   2132: 'Carrier 33 Drive: Error internal communications', class No Acknowledgement, trigger "DB302_HMI_Faults_Carrier33_Faults_1" bit 3
   2133: 'Carrier 33 Drive: Motor overtemperature', class No Acknowledgement, trigger "DB302_HMI_Faults_Carrier33_Faults_1" bit 4
   2134: 'Carrier 33 Drive: Motor overcurrent', class No Acknowledgement, trigger "DB302_HMI_Faults_Carrier33_Faults_1" bit 5
   2135: 'Carrier 33 Drive: Infeed or power unit not ready', class No Acknowledgement, trigger "DB302_HMI_Faults_Carrier33_Faults_1" bit 6
   2136: 'Carrier 33 Drive: Short-circuit/ground fault detected', class No Acknowledgement, trigger "DB302_HMI_Faults_Carrier33_Faults_1" bit 7
   2137: 'Carrier 33 Drive: PROFINET Setpoint timeout', class No Acknowledgement, trigger "DB302_HMI_Faults_Carrier33_Faults_1" bit 8
   2138: 'Carrier 33 Power unit: Overcurrent', class No Acknowledgement, trigger "DB302_HMI_Faults_Carrier33_Faults_1" bit 9
   2139: 'Carrier 33 Power unit: DC link voltage overvoltage', class No Acknowledgement, trigger "DB302_HMI_Faults_Carrier33_Faults_1" bit 10
   2140: 'Carrier 33 Power unit: DC link voltage undervoltage', class No Acknowledgement, trigger "DB302_HMI_Faults_Carrier33_Faults_1" bit 11
   2141: 'Carrier 33 Power unit: Line phase failure in main circuit', class No Acknowledgement, trigger "DB302_HMI_Faults_Carrier33_Faults_1" bit 12
   2142: 'Carrier 33 Power unit: Phase failure motor cable', class No Acknowledgement, trigger "DB302_HMI_Faults_Carrier33_Faults_1" bit 13
   2143: 'Carrier 33 Power unit: Ground fault', class No Acknowledgement, trigger "DB302_HMI_Faults_Carrier33_Faults_1" bit 14
   2144: 'Spare_Fault_2144', class No Acknowledgement, trigger "DB302_HMI_Faults_Carrier33_Faults_1" bit 15
   2145: 'Carrier 33 Motion Off Fault', class No Acknowledgement, trigger "DB302_HMI_Faults_Carrier33_Faults_2" bit 0
   2146: 'Carrier 33 Motion On Fault', class No Acknowledgement, trigger "DB302_HMI_Faults_Carrier33_Faults_2" bit 1
   2147: 'Carrier 33 Spacing Fault', class No Acknowledgement, trigger "DB302_HMI_Faults_Carrier33_Faults_2" bit 2
   2148: 'Carrier 33 Duplicate Carrier Number Fault', class No Acknowledgement, trigger "DB302_HMI_Faults_Carrier33_Faults_2" bit 3
   2149: 'Spare_Fault_2149', class No Acknowledgement, trigger "DB302_HMI_Faults_Carrier33_Faults_2" bit 4
   2150: 'Spare_Fault_2150', class No Acknowledgement, trigger "DB302_HMI_Faults_Carrier33_Faults_2" bit 5
   2151: 'Spare_Fault_2151', class No Acknowledgement, trigger "DB302_HMI_Faults_Carrier33_Faults_2" bit 6
   2152: 'Spare_Fault_2152', class No Acknowledgement, trigger "DB302_HMI_Faults_Carrier33_Faults_2" bit 7
   2153: 'Spare_Fault_2153', class No Acknowledgement, trigger "DB302_HMI_Faults_Carrier33_Faults_2" bit 8
   2154: 'Spare_Fault_2154', class No Acknowledgement, trigger "DB302_HMI_Faults_Carrier33_Faults_2" bit 9
   2155: 'Spare_Fault_2155', class No Acknowledgement, trigger "DB302_HMI_Faults_Carrier33_Faults_2" bit 10
   2156: 'Spare_Fault_2156', class No Acknowledgement, trigger "DB302_HMI_Faults_Carrier33_Faults_2" bit 11
   2157: 'Spare_Fault_2157', class No Acknowledgement, trigger "DB302_HMI_Faults_Carrier33_Faults_2" bit 12
   2158: 'Spare_Fault_2158', class No Acknowledgement, trigger "DB302_HMI_Faults_Carrier33_Faults_2" bit 13
   2159: 'Spare_Fault_2159', class No Acknowledgement, trigger "DB302_HMI_Faults_Carrier33_Faults_2" bit 14
   2160: 'Spare_Fault_2160', class No Acknowledgement, trigger "DB302_HMI_Faults_Carrier33_Faults_2" bit 15
   2161: 'Spare_Fault_2161', class No Acknowledgement, trigger "DB302_HMI_Faults_Carrier33_Faults_3" bit 0
   2162: 'Spare_Fault_2162', class No Acknowledgement, trigger "DB302_HMI_Faults_Carrier33_Faults_3" bit 1
   2163: 'Spare_Fault_2163', class No Acknowledgement, trigger "DB302_HMI_Faults_Carrier33_Faults_3" bit 2
   2164: 'Spare_Fault_2164', class No Acknowledgement, trigger "DB302_HMI_Faults_Carrier33_Faults_3" bit 3
   2165: 'Spare_Fault_2165', class No Acknowledgement, trigger "DB302_HMI_Faults_Carrier33_Faults_3" bit 4
   2166: 'Spare_Fault_2166', class No Acknowledgement, trigger "DB302_HMI_Faults_Carrier33_Faults_3" bit 5
   2167: 'Spare_Fault_2167', class No Acknowledgement, trigger "DB302_HMI_Faults_Carrier33_Faults_3" bit 6
   2168: 'Spare_Fault_2168', class No Acknowledgement, trigger "DB302_HMI_Faults_Carrier33_Faults_3" bit 7
   2169: 'Spare_Fault_2169', class No Acknowledgement, trigger "DB302_HMI_Faults_Carrier33_Faults_3" bit 8
   2170: 'Spare_Fault_2170', class No Acknowledgement, trigger "DB302_HMI_Faults_Carrier33_Faults_3" bit 9
   2171: 'Spare_Fault_2171', class No Acknowledgement, trigger "DB302_HMI_Faults_Carrier33_Faults_3" bit 10
   2172: 'Spare_Fault_2172', class No Acknowledgement, trigger "DB302_HMI_Faults_Carrier33_Faults_3" bit 11
   2173: 'Spare_Fault_2173', class No Acknowledgement, trigger "DB302_HMI_Faults_Carrier33_Faults_3" bit 12
   2174: 'Spare_Fault_2174', class No Acknowledgement, trigger "DB302_HMI_Faults_Carrier33_Faults_3" bit 13
   2175: 'Spare_Fault_2175', class No Acknowledgement, trigger "DB302_HMI_Faults_Carrier33_Faults_3" bit 14
   2176: 'Spare_Fault_2176', class No Acknowledgement, trigger "DB302_HMI_Faults_Carrier33_Faults_3" bit 15
   2177: 'Carrier 34 Disconnect Open Power Fault DI11.0', class No Acknowledgement, trigger "DB302_HMI_Faults_Carrier34_Faults_0" bit 0
   2178: 'Carrier 34 Drive Profinet Comm Fault', class No Acknowledgement, trigger "DB302_HMI_Faults_Carrier34_Faults_0" bit 1
   2179: 'Carrier 34 Production Stop Not Reset', class No Acknowledgement, trigger "DB302_HMI_Faults_Carrier34_Faults_0" bit 2
   2180: 'Carrier 34 CB02122 Tripped', class No Acknowledgement, trigger "DB302_HMI_Faults_Carrier34_Faults_0" bit 3
   2181: 'Carrier 34 CB02123 Tripped', class No Acknowledgement, trigger "DB302_HMI_Faults_Carrier34_Faults_0" bit 4
   2182: 'Carrier 34 AUX1 CB Tripped', class No Acknowledgement, trigger "DB302_HMI_Faults_Carrier34_Faults_0" bit 5
   2183: 'Carrier 34 AUX2 CB Tripped', class No Acknowledgement, trigger "DB302_HMI_Faults_Carrier34_Faults_0" bit 6
   2184: 'Carrier 34 PLC Not Communicating', class No Acknowledgement, trigger "DB302_HMI_Faults_Carrier34_Faults_0" bit 7
   2185: 'Carrier 34 Safe Input Card Fault', class No Acknowledgement, trigger "DB302_HMI_Faults_Carrier34_Faults_0" bit 8
   2186: 'Carrier 34 Safe Output Card Fault', class No Acknowledgement, trigger "DB302_HMI_Faults_Carrier34_Faults_0" bit 9
   2187: 'Carrier 34 Standard Input Card Fault', class No Acknowledgement, trigger "DB302_HMI_Faults_Carrier34_Faults_0" bit 10
   2188: 'Carrier 34 Standard Output Card Fault', class No Acknowledgement, trigger "DB302_HMI_Faults_Carrier34_Faults_0" bit 11
   2189: 'Carrier 34 Encoder Position Fault', class No Acknowledgement, trigger "DB302_HMI_Faults_Carrier34_Faults_0" bit 12
   2190: 'Carrier 34 Encoder Internal Error', class No Acknowledgement, trigger "DB302_HMI_Faults_Carrier34_Faults_0" bit 13
   2191: 'Carrier 34 Encoder Comm Fault', class No Acknowledgement, trigger "DB302_HMI_Faults_Carrier34_Faults_0" bit 14
   2192: 'Carrier 34 HMI Comm Fault', class No Acknowledgement, trigger "DB302_HMI_Faults_Carrier34_Faults_0" bit 15
   2193: 'Carrier 34 Crash Detection Fault', class No Acknowledgement, trigger "DB302_HMI_Faults_Carrier34_Faults_1" bit 0
   2194: 'Carrier 34 Carrier Number Invalid', class No Acknowledgement, trigger "DB302_HMI_Faults_Carrier34_Faults_1" bit 1
   2195: 'Carrier 34 Drive: PROFINET configuration error', class No Acknowledgement, trigger "DB302_HMI_Faults_Carrier34_Faults_1" bit 2
   2196: 'Carrier 34 Drive: Error internal communications', class No Acknowledgement, trigger "DB302_HMI_Faults_Carrier34_Faults_1" bit 3
   2197: 'Carrier 34 Drive: Motor overtemperature', class No Acknowledgement, trigger "DB302_HMI_Faults_Carrier34_Faults_1" bit 4
   2198: 'Carrier 34 Drive: Motor overcurrent', class No Acknowledgement, trigger "DB302_HMI_Faults_Carrier34_Faults_1" bit 5
   2199: 'Carrier 34 Drive: Infeed or power unit not ready', class No Acknowledgement, trigger "DB302_HMI_Faults_Carrier34_Faults_1" bit 6
   2200: 'Carrier 34 Drive: Short-circuit/ground fault detected', class No Acknowledgement, trigger "DB302_HMI_Faults_Carrier34_Faults_1" bit 7
   2201: 'Carrier 34 Drive: PROFINET Setpoint timeout', class No Acknowledgement, trigger "DB302_HMI_Faults_Carrier34_Faults_1" bit 8
   2202: 'Carrier 34 Power unit: Overcurrent', class No Acknowledgement, trigger "DB302_HMI_Faults_Carrier34_Faults_1" bit 9
   2203: 'Carrier 34 Power unit: DC link voltage overvoltage', class No Acknowledgement, trigger "DB302_HMI_Faults_Carrier34_Faults_1" bit 10
   2204: 'Carrier 34 Power unit: DC link voltage undervoltage', class No Acknowledgement, trigger "DB302_HMI_Faults_Carrier34_Faults_1" bit 11
   2205: 'Carrier 34 Power unit: Line phase failure in main circuit', class No Acknowledgement, trigger "DB302_HMI_Faults_Carrier34_Faults_1" bit 12
   2206: 'Carrier 34 Power unit: Phase failure motor cable', class No Acknowledgement, trigger "DB302_HMI_Faults_Carrier34_Faults_1" bit 13
   2207: 'Carrier 34 Power unit: Ground fault', class No Acknowledgement, trigger "DB302_HMI_Faults_Carrier34_Faults_1" bit 14
   2208: 'Spare_Fault_2208', class No Acknowledgement, trigger "DB302_HMI_Faults_Carrier34_Faults_1" bit 15
   2209: 'Carrier 34 Motion Off Fault', class No Acknowledgement, trigger "DB302_HMI_Faults_Carrier34_Faults_2" bit 0
   2210: 'Carrier 34 Motion On Fault', class No Acknowledgement, trigger "DB302_HMI_Faults_Carrier34_Faults_2" bit 1
   2211: 'Carrier 34 Spacing Fault', class No Acknowledgement, trigger "DB302_HMI_Faults_Carrier34_Faults_2" bit 2
   2212: 'Carrier 34 Duplicate Carrier Number Fault', class No Acknowledgement, trigger "DB302_HMI_Faults_Carrier34_Faults_2" bit 3
   2213: 'Spare_Fault_2213', class No Acknowledgement, trigger "DB302_HMI_Faults_Carrier34_Faults_2" bit 4
   2214: 'Spare_Fault_2214', class No Acknowledgement, trigger "DB302_HMI_Faults_Carrier34_Faults_2" bit 5
   2215: 'Spare_Fault_2215', class No Acknowledgement, trigger "DB302_HMI_Faults_Carrier34_Faults_2" bit 6
   2216: 'Spare_Fault_2216', class No Acknowledgement, trigger "DB302_HMI_Faults_Carrier34_Faults_2" bit 7
   2217: 'Spare_Fault_2217', class No Acknowledgement, trigger "DB302_HMI_Faults_Carrier34_Faults_2" bit 8
   2218: 'Spare_Fault_2218', class No Acknowledgement, trigger "DB302_HMI_Faults_Carrier34_Faults_2" bit 9
   2219: 'Spare_Fault_2219', class No Acknowledgement, trigger "DB302_HMI_Faults_Carrier34_Faults_2" bit 10
   2220: 'Spare_Fault_2220', class No Acknowledgement, trigger "DB302_HMI_Faults_Carrier34_Faults_2" bit 11
   2221: 'Spare_Fault_2221', class No Acknowledgement, trigger "DB302_HMI_Faults_Carrier34_Faults_2" bit 12
   2222: 'Spare_Fault_2222', class No Acknowledgement, trigger "DB302_HMI_Faults_Carrier34_Faults_2" bit 13
   2223: 'Spare_Fault_2223', class No Acknowledgement, trigger "DB302_HMI_Faults_Carrier34_Faults_2" bit 14
   2224: 'Spare_Fault_2224', class No Acknowledgement, trigger "DB302_HMI_Faults_Carrier34_Faults_2" bit 15
   2225: 'Spare_Fault_2225', class No Acknowledgement, trigger "DB302_HMI_Faults_Carrier34_Faults_3" bit 0
   2226: 'Spare_Fault_2226', class No Acknowledgement, trigger "DB302_HMI_Faults_Carrier34_Faults_3" bit 1
   2227: 'Spare_Fault_2227', class No Acknowledgement, trigger "DB302_HMI_Faults_Carrier34_Faults_3" bit 2
   2228: 'Spare_Fault_2228', class No Acknowledgement, trigger "DB302_HMI_Faults_Carrier34_Faults_3" bit 3
   2229: 'Spare_Fault_2229', class No Acknowledgement, trigger "DB302_HMI_Faults_Carrier34_Faults_3" bit 4
   2230: 'Spare_Fault_2230', class No Acknowledgement, trigger "DB302_HMI_Faults_Carrier34_Faults_3" bit 5
   2231: 'Spare_Fault_2231', class No Acknowledgement, trigger "DB302_HMI_Faults_Carrier34_Faults_3" bit 6
   2232: 'Spare_Fault_2232', class No Acknowledgement, trigger "DB302_HMI_Faults_Carrier34_Faults_3" bit 7
   2233: 'Spare_Fault_2233', class No Acknowledgement, trigger "DB302_HMI_Faults_Carrier34_Faults_3" bit 8
   2234: 'Spare_Fault_2234', class No Acknowledgement, trigger "DB302_HMI_Faults_Carrier34_Faults_3" bit 9
   2235: 'Spare_Fault_2235', class No Acknowledgement, trigger "DB302_HMI_Faults_Carrier34_Faults_3" bit 10
   2236: 'Spare_Fault_2236', class No Acknowledgement, trigger "DB302_HMI_Faults_Carrier34_Faults_3" bit 11
   2237: 'Spare_Fault_2237', class No Acknowledgement, trigger "DB302_HMI_Faults_Carrier34_Faults_3" bit 12
   2238: 'Spare_Fault_2238', class No Acknowledgement, trigger "DB302_HMI_Faults_Carrier34_Faults_3" bit 13
   2239: 'Spare_Fault_2239', class No Acknowledgement, trigger "DB302_HMI_Faults_Carrier34_Faults_3" bit 14
   2240: 'Spare_Fault_2240', class No Acknowledgement, trigger "DB302_HMI_Faults_Carrier34_Faults_3" bit 15
   2241: 'Carrier 35 Disconnect Open Power Fault DI11.0', class No Acknowledgement, trigger "DB302_HMI_Faults_Carrier35_Faults_0" bit 0
   2242: 'Carrier 35 Drive Profinet Comm Fault', class No Acknowledgement, trigger "DB302_HMI_Faults_Carrier35_Faults_0" bit 1
   2243: 'Carrier 35 Production Stop Not Reset', class No Acknowledgement, trigger "DB302_HMI_Faults_Carrier35_Faults_0" bit 2
   2244: 'Carrier 35 CB02122 Tripped', class No Acknowledgement, trigger "DB302_HMI_Faults_Carrier35_Faults_0" bit 3
   2245: 'Carrier 35 CB02123 Tripped', class No Acknowledgement, trigger "DB302_HMI_Faults_Carrier35_Faults_0" bit 4
   2246: 'Carrier 35 AUX1 CB Tripped', class No Acknowledgement, trigger "DB302_HMI_Faults_Carrier35_Faults_0" bit 5
   2247: 'Carrier 35 AUX2 CB Tripped', class No Acknowledgement, trigger "DB302_HMI_Faults_Carrier35_Faults_0" bit 6
   2248: 'Carrier 35 PLC Not Communicating', class No Acknowledgement, trigger "DB302_HMI_Faults_Carrier35_Faults_0" bit 7
   2249: 'Carrier 35 Safe Input Card Fault', class No Acknowledgement, trigger "DB302_HMI_Faults_Carrier35_Faults_0" bit 8
   2250: 'Carrier 35 Safe Output Card Fault', class No Acknowledgement, trigger "DB302_HMI_Faults_Carrier35_Faults_0" bit 9
   2251: 'Carrier 35 Standard Input Card Fault', class No Acknowledgement, trigger "DB302_HMI_Faults_Carrier35_Faults_0" bit 10
   2252: 'Carrier 35 Standard Output Card Fault', class No Acknowledgement, trigger "DB302_HMI_Faults_Carrier35_Faults_0" bit 11
   2253: 'Carrier 35 Encoder Position Fault', class No Acknowledgement, trigger "DB302_HMI_Faults_Carrier35_Faults_0" bit 12
   2254: 'Carrier 35 Encoder Internal Error', class No Acknowledgement, trigger "DB302_HMI_Faults_Carrier35_Faults_0" bit 13
   2255: 'Carrier 35 Encoder Comm Fault', class No Acknowledgement, trigger "DB302_HMI_Faults_Carrier35_Faults_0" bit 14
   2256: 'Carrier 35 HMI Comm Fault', class No Acknowledgement, trigger "DB302_HMI_Faults_Carrier35_Faults_0" bit 15
   2257: 'Carrier 35 Crash Detection Fault', class No Acknowledgement, trigger "DB302_HMI_Faults_Carrier35_Faults_1" bit 0
   2258: 'Carrier 35 Carrier Number Invalid', class No Acknowledgement, trigger "DB302_HMI_Faults_Carrier35_Faults_1" bit 1
   2259: 'Carrier 35 Drive: PROFINET configuration error', class No Acknowledgement, trigger "DB302_HMI_Faults_Carrier35_Faults_1" bit 2
   2260: 'Carrier 35 Drive: Error internal communications', class No Acknowledgement, trigger "DB302_HMI_Faults_Carrier35_Faults_1" bit 3
   2261: 'Carrier 35 Drive: Motor overtemperature', class No Acknowledgement, trigger "DB302_HMI_Faults_Carrier35_Faults_1" bit 4
   2262: 'Carrier 35 Drive: Motor overcurrent', class No Acknowledgement, trigger "DB302_HMI_Faults_Carrier35_Faults_1" bit 5
   2263: 'Carrier 35 Drive: Infeed or power unit not ready', class No Acknowledgement, trigger "DB302_HMI_Faults_Carrier35_Faults_1" bit 6
   2264: 'Carrier 35 Drive: Short-circuit/ground fault detected', class No Acknowledgement, trigger "DB302_HMI_Faults_Carrier35_Faults_1" bit 7
   2265: 'Carrier 35 Drive: PROFINET Setpoint timeout', class No Acknowledgement, trigger "DB302_HMI_Faults_Carrier35_Faults_1" bit 8
   2266: 'Carrier 35 Power unit: Overcurrent', class No Acknowledgement, trigger "DB302_HMI_Faults_Carrier35_Faults_1" bit 9
   2267: 'Carrier 35 Power unit: DC link voltage overvoltage', class No Acknowledgement, trigger "DB302_HMI_Faults_Carrier35_Faults_1" bit 10
   2268: 'Carrier 35 Power unit: DC link voltage undervoltage', class No Acknowledgement, trigger "DB302_HMI_Faults_Carrier35_Faults_1" bit 11
   2269: 'Carrier 35 Power unit: Line phase failure in main circuit', class No Acknowledgement, trigger "DB302_HMI_Faults_Carrier35_Faults_1" bit 12
   2270: 'Carrier 35 Power unit: Phase failure motor cable', class No Acknowledgement, trigger "DB302_HMI_Faults_Carrier35_Faults_1" bit 13
   2271: 'Carrier 35 Power unit: Ground fault', class No Acknowledgement, trigger "DB302_HMI_Faults_Carrier35_Faults_1" bit 14
   2272: 'Spare_Fault_2272', class No Acknowledgement, trigger "DB302_HMI_Faults_Carrier35_Faults_1" bit 15
   2273: 'Carrier 35 Motion Off Fault', class No Acknowledgement, trigger "DB302_HMI_Faults_Carrier35_Faults_2" bit 0
   2274: 'Carrier 35 Motion On Fault', class No Acknowledgement, trigger "DB302_HMI_Faults_Carrier35_Faults_2" bit 1
   2275: 'Carrier 35 Spacing Fault', class No Acknowledgement, trigger "DB302_HMI_Faults_Carrier35_Faults_2" bit 2
   2276: 'Carrier 35 Duplicate Carrier Number Fault', class No Acknowledgement, trigger "DB302_HMI_Faults_Carrier35_Faults_2" bit 3
   2277: 'Spare_Fault_2277', class No Acknowledgement, trigger "DB302_HMI_Faults_Carrier35_Faults_2" bit 4
   2278: 'Spare_Fault_2278', class No Acknowledgement, trigger "DB302_HMI_Faults_Carrier35_Faults_2" bit 5
   2279: 'Spare_Fault_2279', class No Acknowledgement, trigger "DB302_HMI_Faults_Carrier35_Faults_2" bit 6
   2280: 'Spare_Fault_2280', class No Acknowledgement, trigger "DB302_HMI_Faults_Carrier35_Faults_2" bit 7
   2281: 'Spare_Fault_2281', class No Acknowledgement, trigger "DB302_HMI_Faults_Carrier35_Faults_2" bit 8
   2282: 'Spare_Fault_2282', class No Acknowledgement, trigger "DB302_HMI_Faults_Carrier35_Faults_2" bit 9
   2283: 'Spare_Fault_2283', class No Acknowledgement, trigger "DB302_HMI_Faults_Carrier35_Faults_2" bit 10
   2284: 'Spare_Fault_2284', class No Acknowledgement, trigger "DB302_HMI_Faults_Carrier35_Faults_2" bit 11
   2285: 'Spare_Fault_2285', class No Acknowledgement, trigger "DB302_HMI_Faults_Carrier35_Faults_2" bit 12
   2286: 'Spare_Fault_2286', class No Acknowledgement, trigger "DB302_HMI_Faults_Carrier35_Faults_2" bit 13
   2287: 'Spare_Fault_2287', class No Acknowledgement, trigger "DB302_HMI_Faults_Carrier35_Faults_2" bit 14
   2288: 'Spare_Fault_2288', class No Acknowledgement, trigger "DB302_HMI_Faults_Carrier35_Faults_2" bit 15
   2289: 'Spare_Fault_2289', class No Acknowledgement, trigger "DB302_HMI_Faults_Carrier35_Faults_3" bit 0
   2290: 'Spare_Fault_2290', class No Acknowledgement, trigger "DB302_HMI_Faults_Carrier35_Faults_3" bit 1
   2291: 'Spare_Fault_2291', class No Acknowledgement, trigger "DB302_HMI_Faults_Carrier35_Faults_3" bit 2
   2292: 'Spare_Fault_2292', class No Acknowledgement, trigger "DB302_HMI_Faults_Carrier35_Faults_3" bit 3
   2293: 'Spare_Fault_2293', class No Acknowledgement, trigger "DB302_HMI_Faults_Carrier35_Faults_3" bit 4
   2294: 'Spare_Fault_2294', class No Acknowledgement, trigger "DB302_HMI_Faults_Carrier35_Faults_3" bit 5
   2295: 'Spare_Fault_2295', class No Acknowledgement, trigger "DB302_HMI_Faults_Carrier35_Faults_3" bit 6
   2296: 'Spare_Fault_2296', class No Acknowledgement, trigger "DB302_HMI_Faults_Carrier35_Faults_3" bit 7
   2297: 'Spare_Fault_2297', class No Acknowledgement, trigger "DB302_HMI_Faults_Carrier35_Faults_3" bit 8
   2298: 'Spare_Fault_2298', class No Acknowledgement, trigger "DB302_HMI_Faults_Carrier35_Faults_3" bit 9
   2299: 'Spare_Fault_2299', class No Acknowledgement, trigger "DB302_HMI_Faults_Carrier35_Faults_3" bit 10
   2300: 'Spare_Fault_2300', class No Acknowledgement, trigger "DB302_HMI_Faults_Carrier35_Faults_3" bit 11
   2301: 'Spare_Fault_2301', class No Acknowledgement, trigger "DB302_HMI_Faults_Carrier35_Faults_3" bit 12
   2302: 'Spare_Fault_2302', class No Acknowledgement, trigger "DB302_HMI_Faults_Carrier35_Faults_3" bit 13
   2303: 'Spare_Fault_2303', class No Acknowledgement, trigger "DB302_HMI_Faults_Carrier35_Faults_3" bit 14
   2304: 'Spare_Fault_2304', class No Acknowledgement, trigger "DB302_HMI_Faults_Carrier35_Faults_3" bit 15
   2305: 'Carrier36 Disconnect Open Power Fault DI11.0', class No Acknowledgement, trigger "DB302_HMI_Faults_Carrier36_Faults_0" bit 0
   2306: 'Carrier36 Drive Profinet Comm Fault', class No Acknowledgement, trigger "DB302_HMI_Faults_Carrier36_Faults_0" bit 1
   2307: 'Carrier36 Production Stop Not Reset', class No Acknowledgement, trigger "DB302_HMI_Faults_Carrier36_Faults_0" bit 2
   2308: 'Carrier36 CB02122 Tripped', class No Acknowledgement, trigger "DB302_HMI_Faults_Carrier36_Faults_0" bit 3
   2309: 'Carrier36 CB02123 Tripped', class No Acknowledgement, trigger "DB302_HMI_Faults_Carrier36_Faults_0" bit 4
   2310: 'Carrier36 AUX1 CB Tripped', class No Acknowledgement, trigger "DB302_HMI_Faults_Carrier36_Faults_0" bit 5
   2311: 'Carrier36 AUX2 CB Tripped', class No Acknowledgement, trigger "DB302_HMI_Faults_Carrier36_Faults_0" bit 6
   2312: 'Carrier36 PLC Not Communicating', class No Acknowledgement, trigger "DB302_HMI_Faults_Carrier36_Faults_0" bit 7
   2313: 'Carrier36 Safe Input Card Fault', class No Acknowledgement, trigger "DB302_HMI_Faults_Carrier36_Faults_0" bit 8
   2314: 'Carrier36 Safe Output Card Fault', class No Acknowledgement, trigger "DB302_HMI_Faults_Carrier36_Faults_0" bit 9
   2315: 'Carrier36 Standard Input Card Fault', class No Acknowledgement, trigger "DB302_HMI_Faults_Carrier36_Faults_0" bit 10
   2316: 'Carrier36 Standard Output Card Fault', class No Acknowledgement, trigger "DB302_HMI_Faults_Carrier36_Faults_0" bit 11
   2317: 'Carrier36 Encoder Position Fault', class No Acknowledgement, trigger "DB302_HMI_Faults_Carrier36_Faults_0" bit 12
   2318: 'Carrier36 Encoder Internal Error', class No Acknowledgement, trigger "DB302_HMI_Faults_Carrier36_Faults_0" bit 13
   2319: 'Carrier36 Encoder Comm Fault', class No Acknowledgement, trigger "DB302_HMI_Faults_Carrier36_Faults_0" bit 14
   2320: 'Carrier36 HMI Comm Fault', class No Acknowledgement, trigger "DB302_HMI_Faults_Carrier36_Faults_0" bit 15
   2321: 'Carrier36 Crash Detection Fault', class No Acknowledgement, trigger "DB302_HMI_Faults_Carrier36_Faults_1" bit 0
   2322: 'Carrier36 Carrier Number Invalid', class No Acknowledgement, trigger "DB302_HMI_Faults_Carrier36_Faults_1" bit 1
   2323: 'Carrier36 Drive: PROFINET configuration error', class No Acknowledgement, trigger "DB302_HMI_Faults_Carrier36_Faults_1" bit 2
   2324: 'Carrier36 Drive: Error internal communications', class No Acknowledgement, trigger "DB302_HMI_Faults_Carrier36_Faults_1" bit 3
   2325: 'Carrier36 Drive: Motor overtemperature', class No Acknowledgement, trigger "DB302_HMI_Faults_Carrier36_Faults_1" bit 4
   2326: 'Carrier36 Drive: Motor overcurrent', class No Acknowledgement, trigger "DB302_HMI_Faults_Carrier36_Faults_1" bit 5
   2327: 'Carrier36 Drive: Infeed or power unit not ready', class No Acknowledgement, trigger "DB302_HMI_Faults_Carrier36_Faults_1" bit 6
   2328: 'Carrier36 Drive: Short-circuit/ground fault detected', class No Acknowledgement, trigger "DB302_HMI_Faults_Carrier36_Faults_1" bit 7
   2329: 'Carrier36 Drive: PROFINET Setpoint timeout', class No Acknowledgement, trigger "DB302_HMI_Faults_Carrier36_Faults_1" bit 8
   2330: 'Carrier36 Power unit: Overcurrent', class No Acknowledgement, trigger "DB302_HMI_Faults_Carrier36_Faults_1" bit 9
   2331: 'Carrier36 Power unit: DC link voltage overvoltage', class No Acknowledgement, trigger "DB302_HMI_Faults_Carrier36_Faults_1" bit 10
   2332: 'Carrier36 Power unit: DC link voltage undervoltage', class No Acknowledgement, trigger "DB302_HMI_Faults_Carrier36_Faults_1" bit 11
   2333: 'Carrier36 Power unit: Line phase failure in main circuit', class No Acknowledgement, trigger "DB302_HMI_Faults_Carrier36_Faults_1" bit 12
   2334: 'Carrier36 Power unit: Phase failure motor cable', class No Acknowledgement, trigger "DB302_HMI_Faults_Carrier36_Faults_1" bit 13
   2335: 'Carrier36 Power unit: Ground fault', class No Acknowledgement, trigger "DB302_HMI_Faults_Carrier36_Faults_1" bit 14
   2336: 'Spare_Fault_2336', class No Acknowledgement, trigger "DB302_HMI_Faults_Carrier36_Faults_1" bit 15
   2337: 'Carrier36 Motion Off Fault', class No Acknowledgement, trigger "DB302_HMI_Faults_Carrier36_Faults_2" bit 0
   2338: 'Carrier36 Motion On Fault', class No Acknowledgement, trigger "DB302_HMI_Faults_Carrier36_Faults_2" bit 1
   2339: 'Carrier36 Spacing Fault', class No Acknowledgement, trigger "DB302_HMI_Faults_Carrier36_Faults_2" bit 2
   2340: 'Carrier36 Duplicate Carrier Number Fault', class No Acknowledgement, trigger "DB302_HMI_Faults_Carrier36_Faults_2" bit 3
   2341: 'Spare_Fault_2341', class No Acknowledgement, trigger "DB302_HMI_Faults_Carrier36_Faults_2" bit 4
   2342: 'Spare_Fault_2342', class No Acknowledgement, trigger "DB302_HMI_Faults_Carrier36_Faults_2" bit 5
   2343: 'Spare_Fault_2343', class No Acknowledgement, trigger "DB302_HMI_Faults_Carrier36_Faults_2" bit 6
   2344: 'Spare_Fault_2344', class No Acknowledgement, trigger "DB302_HMI_Faults_Carrier36_Faults_2" bit 7
   2345: 'Spare_Fault_2345', class No Acknowledgement, trigger "DB302_HMI_Faults_Carrier36_Faults_2" bit 8
   2346: 'Spare_Fault_2346', class No Acknowledgement, trigger "DB302_HMI_Faults_Carrier36_Faults_2" bit 9
   2347: 'Spare_Fault_2347', class No Acknowledgement, trigger "DB302_HMI_Faults_Carrier36_Faults_2" bit 10
   2348: 'Spare_Fault_2348', class No Acknowledgement, trigger "DB302_HMI_Faults_Carrier36_Faults_2" bit 11
   2349: 'Spare_Fault_2349', class No Acknowledgement, trigger "DB302_HMI_Faults_Carrier36_Faults_2" bit 12
   2350: 'Spare_Fault_2350', class No Acknowledgement, trigger "DB302_HMI_Faults_Carrier36_Faults_2" bit 13
   2351: 'Spare_Fault_2351', class No Acknowledgement, trigger "DB302_HMI_Faults_Carrier36_Faults_2" bit 14
   2352: 'Spare_Fault_2352', class No Acknowledgement, trigger "DB302_HMI_Faults_Carrier36_Faults_2" bit 15
   2353: 'Spare_Fault_2353', class No Acknowledgement, trigger "DB302_HMI_Faults_Carrier36_Faults_3" bit 0
   2354: 'Spare_Fault_2354', class No Acknowledgement, trigger "DB302_HMI_Faults_Carrier36_Faults_3" bit 1
   2355: 'Spare_Fault_2355', class No Acknowledgement, trigger "DB302_HMI_Faults_Carrier36_Faults_3" bit 2
   2356: 'Spare_Fault_2356', class No Acknowledgement, trigger "DB302_HMI_Faults_Carrier36_Faults_3" bit 3
   2357: 'Spare_Fault_2357', class No Acknowledgement, trigger "DB302_HMI_Faults_Carrier36_Faults_3" bit 4
   2358: 'Spare_Fault_2358', class No Acknowledgement, trigger "DB302_HMI_Faults_Carrier36_Faults_3" bit 5
   2359: 'Spare_Fault_2359', class No Acknowledgement, trigger "DB302_HMI_Faults_Carrier36_Faults_3" bit 6
   2360: 'Spare_Fault_2360', class No Acknowledgement, trigger "DB302_HMI_Faults_Carrier36_Faults_3" bit 7
   2361: 'Spare_Fault_2361', class No Acknowledgement, trigger "DB302_HMI_Faults_Carrier36_Faults_3" bit 8
   2362: 'Spare_Fault_2362', class No Acknowledgement, trigger "DB302_HMI_Faults_Carrier36_Faults_3" bit 9
   2363: 'Spare_Fault_2363', class No Acknowledgement, trigger "DB302_HMI_Faults_Carrier36_Faults_3" bit 10
   2364: 'Spare_Fault_2364', class No Acknowledgement, trigger "DB302_HMI_Faults_Carrier36_Faults_3" bit 11
   2365: 'Spare_Fault_2365', class No Acknowledgement, trigger "DB302_HMI_Faults_Carrier36_Faults_3" bit 12
   2366: 'Spare_Fault_2366', class No Acknowledgement, trigger "DB302_HMI_Faults_Carrier36_Faults_3" bit 13
   2367: 'Spare_Fault_2367', class No Acknowledgement, trigger "DB302_HMI_Faults_Carrier36_Faults_3" bit 14
   2368: 'Spare_Fault_2368', class No Acknowledgement, trigger "DB302_HMI_Faults_Carrier36_Faults_3" bit 15
   2369: 'Carrier 37 Disconnect Open Power Fault DI11.0', class No Acknowledgement, trigger "DB302_HMI_Faults_Carrier37_Faults_0" bit 0
   2370: 'Carrier 37 Drive Profinet Comm Fault', class No Acknowledgement, trigger "DB302_HMI_Faults_Carrier37_Faults_0" bit 1
   2371: 'Carrier 37 Production Stop Not Reset', class No Acknowledgement, trigger "DB302_HMI_Faults_Carrier37_Faults_0" bit 2
   2372: 'Carrier 37 CB02122 Tripped', class No Acknowledgement, trigger "DB302_HMI_Faults_Carrier37_Faults_0" bit 3
   2373: 'Carrier 37 CB02123 Tripped', class No Acknowledgement, trigger "DB302_HMI_Faults_Carrier37_Faults_0" bit 4
   2374: 'Carrier 37 AUX1 CB Tripped', class No Acknowledgement, trigger "DB302_HMI_Faults_Carrier37_Faults_0" bit 5
   2375: 'Carrier 37 AUX2 CB Tripped', class No Acknowledgement, trigger "DB302_HMI_Faults_Carrier37_Faults_0" bit 6
   2376: 'Carrier 37 PLC Not Communicating', class No Acknowledgement, trigger "DB302_HMI_Faults_Carrier37_Faults_0" bit 7
   2377: 'Carrier 37 Safe Input Card Fault', class No Acknowledgement, trigger "DB302_HMI_Faults_Carrier37_Faults_0" bit 8
   2378: 'Carrier 37 Safe Output Card Fault', class No Acknowledgement, trigger "DB302_HMI_Faults_Carrier37_Faults_0" bit 9
   2379: 'Carrier 37 Standard Input Card Fault', class No Acknowledgement, trigger "DB302_HMI_Faults_Carrier37_Faults_0" bit 10
   2380: 'Carrier 37 Standard Output Card Fault', class No Acknowledgement, trigger "DB302_HMI_Faults_Carrier37_Faults_0" bit 11
   2381: 'Carrier 37 Encoder Position Fault', class No Acknowledgement, trigger "DB302_HMI_Faults_Carrier37_Faults_0" bit 12
   2382: 'Carrier 37 Encoder Internal Error', class No Acknowledgement, trigger "DB302_HMI_Faults_Carrier37_Faults_0" bit 13
   2383: 'Carrier 37 Encoder Comm Fault', class No Acknowledgement, trigger "DB302_HMI_Faults_Carrier37_Faults_0" bit 14
   2384: 'Carrier 37 HMI Comm Fault', class No Acknowledgement, trigger "DB302_HMI_Faults_Carrier37_Faults_0" bit 15
   2385: 'Carrier 37 Crash Detection Fault', class No Acknowledgement, trigger "DB302_HMI_Faults_Carrier37_Faults_1" bit 0
   2386: 'Carrier 37 Carrier Number Invalid', class No Acknowledgement, trigger "DB302_HMI_Faults_Carrier37_Faults_1" bit 1
   2387: 'Carrier 37 Drive: PROFINET configuration error', class No Acknowledgement, trigger "DB302_HMI_Faults_Carrier37_Faults_1" bit 2
   2388: 'Carrier 37 Drive: Error internal communications', class No Acknowledgement, trigger "DB302_HMI_Faults_Carrier37_Faults_1" bit 3
   2389: 'Carrier 37 Drive: Motor overtemperature', class No Acknowledgement, trigger "DB302_HMI_Faults_Carrier37_Faults_1" bit 4
   2390: 'Carrier 37 Drive: Motor overcurrent', class No Acknowledgement, trigger "DB302_HMI_Faults_Carrier37_Faults_1" bit 5
   2391: 'Carrier 37 Drive: Infeed or power unit not ready', class No Acknowledgement, trigger "DB302_HMI_Faults_Carrier37_Faults_1" bit 6
   2392: 'Carrier 37 Drive: Short-circuit/ground fault detected', class No Acknowledgement, trigger "DB302_HMI_Faults_Carrier37_Faults_1" bit 7
   2393: 'Carrier 37 Drive: PROFINET Setpoint timeout', class No Acknowledgement, trigger "DB302_HMI_Faults_Carrier37_Faults_1" bit 8
   2394: 'Carrier 37 Power unit: Overcurrent', class No Acknowledgement, trigger "DB302_HMI_Faults_Carrier37_Faults_1" bit 9
   2395: 'Carrier 37 Power unit: DC link voltage overvoltage', class No Acknowledgement, trigger "DB302_HMI_Faults_Carrier37_Faults_1" bit 10
   2396: 'Carrier 37 Power unit: DC link voltage undervoltage', class No Acknowledgement, trigger "DB302_HMI_Faults_Carrier37_Faults_1" bit 11
   2397: 'Carrier 37 Power unit: Line phase failure in main circuit', class No Acknowledgement, trigger "DB302_HMI_Faults_Carrier37_Faults_1" bit 12
   2398: 'Carrier 37 Power unit: Phase failure motor cable', class No Acknowledgement, trigger "DB302_HMI_Faults_Carrier37_Faults_1" bit 13
   2399: 'Carrier 37 Power unit: Ground fault', class No Acknowledgement, trigger "DB302_HMI_Faults_Carrier37_Faults_1" bit 14
   2400: 'Spare_Fault_2400', class No Acknowledgement, trigger "DB302_HMI_Faults_Carrier37_Faults_1" bit 15
   2401: 'Carrier 37 Motion Off Fault', class No Acknowledgement, trigger "DB302_HMI_Faults_Carrier37_Faults_2" bit 0
   2402: 'Carrier 37 Motion On Fault', class No Acknowledgement, trigger "DB302_HMI_Faults_Carrier37_Faults_2" bit 1
   2403: 'Carrier 37 Spacing Fault', class No Acknowledgement, trigger "DB302_HMI_Faults_Carrier37_Faults_2" bit 2
   2404: 'Carrier 37 Duplicate Carrier Number Fault', class No Acknowledgement, trigger "DB302_HMI_Faults_Carrier37_Faults_2" bit 3
   2405: 'Spare_Fault_2405', class No Acknowledgement, trigger "DB302_HMI_Faults_Carrier37_Faults_2" bit 4
   2406: 'Spare_Fault_2406', class No Acknowledgement, trigger "DB302_HMI_Faults_Carrier37_Faults_2" bit 5
   2407: 'Spare_Fault_2407', class No Acknowledgement, trigger "DB302_HMI_Faults_Carrier37_Faults_2" bit 6
   2408: 'Spare_Fault_2408', class No Acknowledgement, trigger "DB302_HMI_Faults_Carrier37_Faults_2" bit 7
   2409: 'Spare_Fault_2409', class No Acknowledgement, trigger "DB302_HMI_Faults_Carrier37_Faults_2" bit 8
   2410: 'Spare_Fault_2410', class No Acknowledgement, trigger "DB302_HMI_Faults_Carrier37_Faults_2" bit 9
   2411: 'Spare_Fault_2411', class No Acknowledgement, trigger "DB302_HMI_Faults_Carrier37_Faults_2" bit 10
   2412: 'Spare_Fault_2412', class No Acknowledgement, trigger "DB302_HMI_Faults_Carrier37_Faults_2" bit 11
   2413: 'Spare_Fault_2413', class No Acknowledgement, trigger "DB302_HMI_Faults_Carrier37_Faults_2" bit 12
   2414: 'Spare_Fault_2414', class No Acknowledgement, trigger "DB302_HMI_Faults_Carrier37_Faults_2" bit 13
   2415: 'Spare_Fault_2415', class No Acknowledgement, trigger "DB302_HMI_Faults_Carrier37_Faults_2" bit 14
   2416: 'Spare_Fault_2416', class No Acknowledgement, trigger "DB302_HMI_Faults_Carrier37_Faults_2" bit 15
   2417: 'Spare_Fault_2417', class No Acknowledgement, trigger "DB302_HMI_Faults_Carrier37_Faults_3" bit 0
   2418: 'Spare_Fault_2418', class No Acknowledgement, trigger "DB302_HMI_Faults_Carrier37_Faults_3" bit 1
   2419: 'Spare_Fault_2419', class No Acknowledgement, trigger "DB302_HMI_Faults_Carrier37_Faults_3" bit 2
   2420: 'Spare_Fault_2420', class No Acknowledgement, trigger "DB302_HMI_Faults_Carrier37_Faults_3" bit 3
   2421: 'Spare_Fault_2421', class No Acknowledgement, trigger "DB302_HMI_Faults_Carrier37_Faults_3" bit 4
   2422: 'Spare_Fault_2422', class No Acknowledgement, trigger "DB302_HMI_Faults_Carrier37_Faults_3" bit 5
   2423: 'Spare_Fault_2423', class No Acknowledgement, trigger "DB302_HMI_Faults_Carrier37_Faults_3" bit 6
   2424: 'Spare_Fault_2424', class No Acknowledgement, trigger "DB302_HMI_Faults_Carrier37_Faults_3" bit 7
   2425: 'Spare_Fault_2425', class No Acknowledgement, trigger "DB302_HMI_Faults_Carrier37_Faults_3" bit 8
   2426: 'Spare_Fault_2426', class No Acknowledgement, trigger "DB302_HMI_Faults_Carrier37_Faults_3" bit 9
   2427: 'Spare_Fault_2427', class No Acknowledgement, trigger "DB302_HMI_Faults_Carrier37_Faults_3" bit 10
   2428: 'Spare_Fault_2428', class No Acknowledgement, trigger "DB302_HMI_Faults_Carrier37_Faults_3" bit 11
   2429: 'Spare_Fault_2429', class No Acknowledgement, trigger "DB302_HMI_Faults_Carrier37_Faults_3" bit 12
   2430: 'Spare_Fault_2430', class No Acknowledgement, trigger "DB302_HMI_Faults_Carrier37_Faults_3" bit 13
   2431: 'Spare_Fault_2431', class No Acknowledgement, trigger "DB302_HMI_Faults_Carrier37_Faults_3" bit 14
   2432: 'Spare_Fault_2432', class No Acknowledgement, trigger "DB302_HMI_Faults_Carrier37_Faults_3" bit 15
   2433: 'Carrier 38 Disconnect Open Power Fault DI11.0', class No Acknowledgement, trigger "DB302_HMI_Faults_Carrier38_Faults_0" bit 0
   2434: 'Carrier 38 Drive Profinet Comm Fault', class No Acknowledgement, trigger "DB302_HMI_Faults_Carrier38_Faults_0" bit 1
   2435: 'Carrier 38 Production Stop Not Reset', class No Acknowledgement, trigger "DB302_HMI_Faults_Carrier38_Faults_0" bit 2
   2436: 'Carrier 38 CB02122 Tripped', class No Acknowledgement, trigger "DB302_HMI_Faults_Carrier38_Faults_0" bit 3
   2437: 'Carrier 38 CB02123 Tripped', class No Acknowledgement, trigger "DB302_HMI_Faults_Carrier38_Faults_0" bit 4
   2438: 'Carrier 38 AUX1 CB Tripped', class No Acknowledgement, trigger "DB302_HMI_Faults_Carrier38_Faults_0" bit 5
   2439: 'Carrier 38 AUX2 CB Tripped', class No Acknowledgement, trigger "DB302_HMI_Faults_Carrier38_Faults_0" bit 6
   2440: 'Carrier 38 PLC Not Communicating', class No Acknowledgement, trigger "DB302_HMI_Faults_Carrier38_Faults_0" bit 7
   2441: 'Carrier 38 Safe Input Card Fault', class No Acknowledgement, trigger "DB302_HMI_Faults_Carrier38_Faults_0" bit 8
   2442: 'Carrier 38 Safe Output Card Fault', class No Acknowledgement, trigger "DB302_HMI_Faults_Carrier38_Faults_0" bit 9
   2443: 'Carrier 38 Standard Input Card Fault', class No Acknowledgement, trigger "DB302_HMI_Faults_Carrier38_Faults_0" bit 10
   2444: 'Carrier 38 Standard Output Card Fault', class No Acknowledgement, trigger "DB302_HMI_Faults_Carrier38_Faults_0" bit 11
   2445: 'Carrier 38 Encoder Position Fault', class No Acknowledgement, trigger "DB302_HMI_Faults_Carrier38_Faults_0" bit 12
   2446: 'Carrier 38 Encoder Internal Error', class No Acknowledgement, trigger "DB302_HMI_Faults_Carrier38_Faults_0" bit 13
   2447: 'Carrier 38 Encoder Comm Fault', class No Acknowledgement, trigger "DB302_HMI_Faults_Carrier38_Faults_0" bit 14
   2448: 'Carrier 38 HMI Comm Fault', class No Acknowledgement, trigger "DB302_HMI_Faults_Carrier38_Faults_0" bit 15
   2449: 'Carrier 38 Crash Detection Fault', class No Acknowledgement, trigger "DB302_HMI_Faults_Carrier38_Faults_1" bit 0
   2450: 'Carrier 38 Carrier Number Invalid', class No Acknowledgement, trigger "DB302_HMI_Faults_Carrier38_Faults_1" bit 1
   2451: 'Carrier 38 Drive: PROFINET configuration error', class No Acknowledgement, trigger "DB302_HMI_Faults_Carrier38_Faults_1" bit 2
   2452: 'Carrier 38 Drive: Error internal communications', class No Acknowledgement, trigger "DB302_HMI_Faults_Carrier38_Faults_1" bit 3
   2453: 'Carrier 38 Drive: Motor overtemperature', class No Acknowledgement, trigger "DB302_HMI_Faults_Carrier38_Faults_1" bit 4
   2454: 'Carrier 38 Drive: Motor overcurrent', class No Acknowledgement, trigger "DB302_HMI_Faults_Carrier38_Faults_1" bit 5
   2455: 'Carrier 38 Drive: Infeed or power unit not ready', class No Acknowledgement, trigger "DB302_HMI_Faults_Carrier38_Faults_1" bit 6
   2456: 'Carrier 38 Drive: Short-circuit/ground fault detected', class No Acknowledgement, trigger "DB302_HMI_Faults_Carrier38_Faults_1" bit 7
   2457: 'Carrier 38 Drive: PROFINET Setpoint timeout', class No Acknowledgement, trigger "DB302_HMI_Faults_Carrier38_Faults_1" bit 8
   2458: 'Carrier 38 Power unit: Overcurrent', class No Acknowledgement, trigger "DB302_HMI_Faults_Carrier38_Faults_1" bit 9
   2459: 'Carrier 38 Power unit: DC link voltage overvoltage', class No Acknowledgement, trigger "DB302_HMI_Faults_Carrier38_Faults_1" bit 10
   2460: 'Carrier 38 Power unit: DC link voltage undervoltage', class No Acknowledgement, trigger "DB302_HMI_Faults_Carrier38_Faults_1" bit 11
   2461: 'Carrier 38 Power unit: Line phase failure in main circuit', class No Acknowledgement, trigger "DB302_HMI_Faults_Carrier38_Faults_1" bit 12
   2462: 'Carrier 38 Power unit: Phase failure motor cable', class No Acknowledgement, trigger "DB302_HMI_Faults_Carrier38_Faults_1" bit 13
   2463: 'Carrier 38 Power unit: Ground fault', class No Acknowledgement, trigger "DB302_HMI_Faults_Carrier38_Faults_1" bit 14
   2464: 'Spare_Fault_2464', class No Acknowledgement, trigger "DB302_HMI_Faults_Carrier38_Faults_1" bit 15
   2465: 'Carrier 38 Motion Off Fault', class No Acknowledgement, trigger "DB302_HMI_Faults_Carrier38_Faults_2" bit 0
   2466: 'Carrier 38 Motion On Fault', class No Acknowledgement, trigger "DB302_HMI_Faults_Carrier38_Faults_2" bit 1
   2467: 'Carrier 38 Spacing Fault', class No Acknowledgement, trigger "DB302_HMI_Faults_Carrier38_Faults_2" bit 2
   2468: 'Carrier 38 Duplicate Carrier Number Fault', class No Acknowledgement, trigger "DB302_HMI_Faults_Carrier38_Faults_2" bit 3
   2469: 'Spare_Fault_2469', class No Acknowledgement, trigger "DB302_HMI_Faults_Carrier38_Faults_2" bit 4
   2470: 'Spare_Fault_2470', class No Acknowledgement, trigger "DB302_HMI_Faults_Carrier38_Faults_2" bit 5
   2471: 'Spare_Fault_2471', class No Acknowledgement, trigger "DB302_HMI_Faults_Carrier38_Faults_2" bit 6
   2472: 'Spare_Fault_2472', class No Acknowledgement, trigger "DB302_HMI_Faults_Carrier38_Faults_2" bit 7
   2473: 'Spare_Fault_2473', class No Acknowledgement, trigger "DB302_HMI_Faults_Carrier38_Faults_2" bit 8
   2474: 'Spare_Fault_2474', class No Acknowledgement, trigger "DB302_HMI_Faults_Carrier38_Faults_2" bit 9
   2475: 'Spare_Fault_2475', class No Acknowledgement, trigger "DB302_HMI_Faults_Carrier38_Faults_2" bit 10
   2476: 'Spare_Fault_2476', class No Acknowledgement, trigger "DB302_HMI_Faults_Carrier38_Faults_2" bit 11
   2477: 'Spare_Fault_2477', class No Acknowledgement, trigger "DB302_HMI_Faults_Carrier38_Faults_2" bit 12
   2478: 'Spare_Fault_2478', class No Acknowledgement, trigger "DB302_HMI_Faults_Carrier38_Faults_2" bit 13
   2479: 'Spare_Fault_2479', class No Acknowledgement, trigger "DB302_HMI_Faults_Carrier38_Faults_2" bit 14
   2480: 'Spare_Fault_2480', class No Acknowledgement, trigger "DB302_HMI_Faults_Carrier38_Faults_2" bit 15
   2481: 'Spare_Fault_2481', class No Acknowledgement, trigger "DB302_HMI_Faults_Carrier38_Faults_3" bit 0
   2482: 'Spare_Fault_2482', class No Acknowledgement, trigger "DB302_HMI_Faults_Carrier38_Faults_3" bit 1
   2483: 'Spare_Fault_2483', class No Acknowledgement, trigger "DB302_HMI_Faults_Carrier38_Faults_3" bit 2
   2484: 'Spare_Fault_2484', class No Acknowledgement, trigger "DB302_HMI_Faults_Carrier38_Faults_3" bit 3
   2485: 'Spare_Fault_2485', class No Acknowledgement, trigger "DB302_HMI_Faults_Carrier38_Faults_3" bit 4
   2486: 'Spare_Fault_2486', class No Acknowledgement, trigger "DB302_HMI_Faults_Carrier38_Faults_3" bit 5
   2487: 'Spare_Fault_2487', class No Acknowledgement, trigger "DB302_HMI_Faults_Carrier38_Faults_3" bit 6
   2488: 'Spare_Fault_2488', class No Acknowledgement, trigger "DB302_HMI_Faults_Carrier38_Faults_3" bit 7
   2489: 'Spare_Fault_2489', class No Acknowledgement, trigger "DB302_HMI_Faults_Carrier38_Faults_3" bit 8
   2490: 'Spare_Fault_2490', class No Acknowledgement, trigger "DB302_HMI_Faults_Carrier38_Faults_3" bit 9
   2491: 'Spare_Fault_2491', class No Acknowledgement, trigger "DB302_HMI_Faults_Carrier38_Faults_3" bit 10
   2492: 'Spare_Fault_2492', class No Acknowledgement, trigger "DB302_HMI_Faults_Carrier38_Faults_3" bit 11
   2493: 'Spare_Fault_2493', class No Acknowledgement, trigger "DB302_HMI_Faults_Carrier38_Faults_3" bit 12
   2494: 'Spare_Fault_2494', class No Acknowledgement, trigger "DB302_HMI_Faults_Carrier38_Faults_3" bit 13
   2495: 'Spare_Fault_2495', class No Acknowledgement, trigger "DB302_HMI_Faults_Carrier38_Faults_3" bit 14
   2496: 'Spare_Fault_2496', class No Acknowledgement, trigger "DB302_HMI_Faults_Carrier38_Faults_3" bit 15
   2497: 'Carrier 39 Disconnect Open Power Fault DI11.0', class No Acknowledgement, trigger "DB302_HMI_Faults_Carrier39_Faults_0" bit 0
   2498: 'Carrier 39 Drive Profinet Comm Fault', class No Acknowledgement, trigger "DB302_HMI_Faults_Carrier39_Faults_0" bit 1
   2499: 'Carrier 39 Production Stop Not Reset', class No Acknowledgement, trigger "DB302_HMI_Faults_Carrier39_Faults_0" bit 2
   2500: 'Carrier 39 CB02122 Tripped', class No Acknowledgement, trigger "DB302_HMI_Faults_Carrier39_Faults_0" bit 3
   2501: 'Carrier 39 CB02123 Tripped', class No Acknowledgement, trigger "DB302_HMI_Faults_Carrier39_Faults_0" bit 4
   2502: 'Carrier 39 AUX1 CB Tripped', class No Acknowledgement, trigger "DB302_HMI_Faults_Carrier39_Faults_0" bit 5
   2503: 'Carrier 39 AUX2 CB Tripped', class No Acknowledgement, trigger "DB302_HMI_Faults_Carrier39_Faults_0" bit 6
   2504: 'Carrier 39 PLC Not Communicating', class No Acknowledgement, trigger "DB302_HMI_Faults_Carrier39_Faults_0" bit 7
   2505: 'Carrier 39 Safe Input Card Fault', class No Acknowledgement, trigger "DB302_HMI_Faults_Carrier39_Faults_0" bit 8
   2506: 'Carrier 39 Safe Output Card Fault', class No Acknowledgement, trigger "DB302_HMI_Faults_Carrier39_Faults_0" bit 9
   2507: 'Carrier 39 Standard Input Card Fault', class No Acknowledgement, trigger "DB302_HMI_Faults_Carrier39_Faults_0" bit 10
   2508: 'Carrier 39 Standard Output Card Fault', class No Acknowledgement, trigger "DB302_HMI_Faults_Carrier39_Faults_0" bit 11
   2509: 'Carrier 39 Encoder Position Fault', class No Acknowledgement, trigger "DB302_HMI_Faults_Carrier39_Faults_0" bit 12
   2510: 'Carrier 39 Encoder Internal Error', class No Acknowledgement, trigger "DB302_HMI_Faults_Carrier39_Faults_0" bit 13
   2511: 'Carrier 39 Encoder Comm Fault', class No Acknowledgement, trigger "DB302_HMI_Faults_Carrier39_Faults_0" bit 14
   2512: 'Carrier 39 HMI Comm Fault', class No Acknowledgement, trigger "DB302_HMI_Faults_Carrier39_Faults_0" bit 15
   2513: 'Carrier 39 Crash Detection Fault', class No Acknowledgement, trigger "DB302_HMI_Faults_Carrier39_Faults_1" bit 0
   2514: 'Carrier 39 Carrier Number Invalid', class No Acknowledgement, trigger "DB302_HMI_Faults_Carrier39_Faults_1" bit 1
   2515: 'Carrier 39 Drive: PROFINET configuration error', class No Acknowledgement, trigger "DB302_HMI_Faults_Carrier39_Faults_1" bit 2
   2516: 'Carrier 39 Drive: Error internal communications', class No Acknowledgement, trigger "DB302_HMI_Faults_Carrier39_Faults_1" bit 3
   2517: 'Carrier 39 Drive: Motor overtemperature', class No Acknowledgement, trigger "DB302_HMI_Faults_Carrier39_Faults_1" bit 4
   2518: 'Carrier 39 Drive: Motor overcurrent', class No Acknowledgement, trigger "DB302_HMI_Faults_Carrier39_Faults_1" bit 5
   2519: 'Carrier 39 Drive: Infeed or power unit not ready', class No Acknowledgement, trigger "DB302_HMI_Faults_Carrier39_Faults_1" bit 6
   2520: 'Carrier 39 Drive: Short-circuit/ground fault detected', class No Acknowledgement, trigger "DB302_HMI_Faults_Carrier39_Faults_1" bit 7
   2521: 'Carrier 39 Drive: PROFINET Setpoint timeout', class No Acknowledgement, trigger "DB302_HMI_Faults_Carrier39_Faults_1" bit 8
   2522: 'Carrier 39 Power unit: Overcurrent', class No Acknowledgement, trigger "DB302_HMI_Faults_Carrier39_Faults_1" bit 9
   2523: 'Carrier 39 Power unit: DC link voltage overvoltage', class No Acknowledgement, trigger "DB302_HMI_Faults_Carrier39_Faults_1" bit 10
   2524: 'Carrier 39 Power unit: DC link voltage undervoltage', class No Acknowledgement, trigger "DB302_HMI_Faults_Carrier39_Faults_1" bit 11
   2525: 'Carrier 39 Power unit: Line phase failure in main circuit', class No Acknowledgement, trigger "DB302_HMI_Faults_Carrier39_Faults_1" bit 12
   2526: 'Carrier 39 Power unit: Phase failure motor cable', class No Acknowledgement, trigger "DB302_HMI_Faults_Carrier39_Faults_1" bit 13
   2527: 'Carrier 39 Power unit: Ground fault', class No Acknowledgement, trigger "DB302_HMI_Faults_Carrier39_Faults_1" bit 14
   2528: 'Spare_Fault_2528', class No Acknowledgement, trigger "DB302_HMI_Faults_Carrier39_Faults_1" bit 15
   2529: 'Carrier 39 Motion Off Fault', class No Acknowledgement, trigger "DB302_HMI_Faults_Carrier39_Faults_2" bit 0
   2530: 'Carrier 39 Motion On Fault', class No Acknowledgement, trigger "DB302_HMI_Faults_Carrier39_Faults_2" bit 1
   2531: 'Carrier 39 Spacing Fault', class No Acknowledgement, trigger "DB302_HMI_Faults_Carrier39_Faults_2" bit 2
   2532: 'Carrier 39 Duplicate Carrier Number Fault', class No Acknowledgement, trigger "DB302_HMI_Faults_Carrier39_Faults_2" bit 3
   2533: 'Spare_Fault_2533', class No Acknowledgement, trigger "DB302_HMI_Faults_Carrier39_Faults_2" bit 4
   2534: 'Spare_Fault_2534', class No Acknowledgement, trigger "DB302_HMI_Faults_Carrier39_Faults_2" bit 5
   2535: 'Spare_Fault_2535', class No Acknowledgement, trigger "DB302_HMI_Faults_Carrier39_Faults_2" bit 6
   2536: 'Spare_Fault_2536', class No Acknowledgement, trigger "DB302_HMI_Faults_Carrier39_Faults_2" bit 7
   2537: 'Spare_Fault_2537', class No Acknowledgement, trigger "DB302_HMI_Faults_Carrier39_Faults_2" bit 8
   2538: 'Spare_Fault_2538', class No Acknowledgement, trigger "DB302_HMI_Faults_Carrier39_Faults_2" bit 9
   2539: 'Spare_Fault_2539', class No Acknowledgement, trigger "DB302_HMI_Faults_Carrier39_Faults_2" bit 10
   2540: 'Spare_Fault_2540', class No Acknowledgement, trigger "DB302_HMI_Faults_Carrier39_Faults_2" bit 11
   2541: 'Spare_Fault_2541', class No Acknowledgement, trigger "DB302_HMI_Faults_Carrier39_Faults_2" bit 12
   2542: 'Spare_Fault_2542', class No Acknowledgement, trigger "DB302_HMI_Faults_Carrier39_Faults_2" bit 13
   2543: 'Spare_Fault_2543', class No Acknowledgement, trigger "DB302_HMI_Faults_Carrier39_Faults_2" bit 14
   2544: 'Spare_Fault_2544', class No Acknowledgement, trigger "DB302_HMI_Faults_Carrier39_Faults_2" bit 15
   2545: 'Spare_Fault_2545', class No Acknowledgement, trigger "DB302_HMI_Faults_Carrier39_Faults_3" bit 0
   2546: 'Spare_Fault_2546', class No Acknowledgement, trigger "DB302_HMI_Faults_Carrier39_Faults_3" bit 1
   2547: 'Spare_Fault_2547', class No Acknowledgement, trigger "DB302_HMI_Faults_Carrier39_Faults_3" bit 2
   2548: 'Spare_Fault_2548', class No Acknowledgement, trigger "DB302_HMI_Faults_Carrier39_Faults_3" bit 3
   2549: 'Spare_Fault_2549', class No Acknowledgement, trigger "DB302_HMI_Faults_Carrier39_Faults_3" bit 4
   2550: 'Spare_Fault_2550', class No Acknowledgement, trigger "DB302_HMI_Faults_Carrier39_Faults_3" bit 5
   2551: 'Spare_Fault_2551', class No Acknowledgement, trigger "DB302_HMI_Faults_Carrier39_Faults_3" bit 6
   2552: 'Spare_Fault_2552', class No Acknowledgement, trigger "DB302_HMI_Faults_Carrier39_Faults_3" bit 7
